// TIA Portal project "YDSLK_HMI_2023-05-10_08-26_V3_00T" (V15.1) (continued)
   "ST_HMI_Var_HMI_r64PositiveAccel_ZouChe_ChuChe" : LReal = PLC ST_HMI_Var.HMI_r64PositiveAccel_ZouChe_ChuChe AT 10-30-00-01-00-21-84-00-13-00, 1 s
   "ST_HMI_Var_HMI_r64AccVelocity_Jog_ChengXing_Up" : LReal = PLC ST_HMI_Var.HMI_r64AccVelocity_Jog_ChengXing_Up AT 10-30-00-01-00-21-84-00-1D-40, 1 s
   "VBS_time_hour" : LReal, internal
   "ST_HMI_Var_HMI_r64Velocity_Jog_JinChe" : LReal = PLC ST_HMI_Var.HMI_r64Velocity_Jog_JinChe AT 10-30-00-01-00-21-84-00-1A-40, 1 s
   "ST_HMI_Var_HMI_alpha_JuanRao_3" : LReal = PLC ST_HMI_Var.HMI_alpha_JuanRao_3 AT 10-30-00-01-00-21-84-00-33-80, 1 s
   "ST_HMI_Var_HMI_r64_LuoSha_Force_DanSha_ZhangLi_FangKai" : LReal = PLC ST_HMI_Var.HMI_r64_LuoSha_Force_DanSha_ZhangLi_FangKai AT 10-30-00-01-00-21-84-00-21-80, 1 s
   "ST_HMI_Var_HMI_r64Height_ShaSui_Start" : LReal = PLC ST_HMI_Var.HMI_r64Height_ShaSui_Start AT 10-30-00-01-00-21-84-00-0A-80, 1 s
   "ST_HMI_Var_HMI_r64Axis_ChengXing_positiveaccelstartjerk_CunRao" : LReal = PLC ST_HMI_Var.HMI_r64Axis_ChengXing_positiveaccelstartjerk_CunRao AT 10-30-00-01-00-21-84-00-3C-80, 1 s
   "ST_HMI_Var_HMI_K_T_M" : LReal = PLC ST_HMI_Var.HMI_K_T_M AT 10-30-00-01-00-21-84-00-43-C0, 1 s
   "ST_HMI_Var_HMI_r64Diameter_ShaGuan_Bottom" : LReal = PLC ST_HMI_Var.HMI_r64Diameter_ShaGuan_Bottom AT 10-30-00-01-00-21-84-00-0C-80, 1 s
   "ST_HMI_Var_HMI_r64Axis_1_ZhangLi_Position_JuanRao_Set_ND" : LReal = PLC ST_HMI_Var.HMI_r64Axis_1_ZhangLi_Position_JuanRao_Set_ND AT 10-30-00-01-00-21-84-00-39-00, 1 s
   "ST_HMI_Var_HMI_r64AccVelocity_Jog_ChuChe" : LReal = PLC ST_HMI_Var.HMI_r64AccVelocity_Jog_ChuChe AT 10-30-00-01-00-21-84-00-1A-00, 1 s
   "ST_HMI_Var_HMI_r64Velocity_Jog_ChengXing_Up" : LReal = PLC ST_HMI_Var.HMI_r64Velocity_Jog_ChengXing_Up AT 10-30-00-01-00-21-84-00-1D-00, 1 s
   "ST_HMI_Var_HMI_cam2_ratio_delt_min" : LReal = PLC ST_HMI_Var.HMI_cam2_ratio_delt_min AT 10-30-00-01-00-21-84-00-30-00, 1 s
   "ST_HMI_Var_HMI_r64Axis_DingZi_Velocity_JuanRao_max" : LReal = PLC ST_HMI_Var.HMI_r64Axis_DingZi_Velocity_JuanRao_max AT 10-30-00-01-00-21-84-00-38-40, 1 s
   "ST_Main_Var_g_bo_Automatic_Running_Status" : Bool = PLC ST_Main_Var.g_bo_Automatic_Running_Status AT 10-01-00-01-00-23-84-00-51-E0, 1 s
   "ST_HMI_Var_HMI_cam_ChengXing_delt_syncoffpositionslave_tuirao" : LReal = PLC ST_HMI_Var.HMI_cam_ChengXing_delt_syncoffpositionslave_tuirao AT 10-30-00-01-00-21-84-00-32-40, 1 s
   "变量_4" : UInt, internal
   "ST_Main_Var_g_r64Axis_DingZi_Velocity_CunRao_ratio" : LReal = PLC ST_Main_Var.g_r64Axis_DingZi_Velocity_CunRao_ratio AT 10-30-00-01-00-23-84-00-32-C0, 1 s
   "变量_2" : WString[10], internal
   "ST_HMI_Var_HMI_r64Axis_ZouChe_negativeaccelstartjerk_JinChe" : LReal = PLC ST_HMI_Var.HMI_r64Axis_ZouChe_negativeaccelstartjerk_JinChe AT 10-30-00-01-00-21-84-00-15-40, 1 s
   "ST_HMI_Var_HMI_r64Axis_1_ZhangLi_Velocity_JuanRao" : LReal = PLC ST_HMI_Var.HMI_r64Axis_1_ZhangLi_Velocity_JuanRao AT 10-30-00-01-00-21-84-00-3B-40, 1 s
   "变量_16" : Bool, internal
   "ST_HMI_Var_HMI_r64_MaoZhou_TouShu" : Int = PLC ST_HMI_Var.HMI_r64_MaoZhou_TouShu AT 10-05-00-01-00-21-84-00-22-00, 1 s
   "ST_HMI_Var_HMI_xit_delt_max" : LReal = PLC ST_HMI_Var.HMI_xit_delt_max AT 10-30-00-01-00-21-84-00-24-00, 1 s
   "ST_HMI_Var_luoshu" : Int = PLC ST_HMI_Var.luoshu AT 10-05-00-01-00-21-84-00-6B-00, 1 s
   "ST_HMI_Var_HMI_r64NianSu_3" : LReal = PLC ST_HMI_Var.HMI_r64NianSu_3 AT 10-30-00-01-00-21-84-00-04-00, 1 s
   "ST_HMI_Var_HMI_boAlarm_NianSuo_PosNon" : Bool = PLC ST_HMI_Var.HMI_boAlarm_NianSuo_PosNon AT 10-01-00-01-00-21-84-00-05-C0, 1 s
   "ST_HMI_Var_HMI_r64NianDu_actual" : LReal = PLC ST_HMI_Var.HMI_r64NianDu_actual AT 10-30-00-01-00-21-84-00-19-40, 1 s
   "ST_HMI_Var_HMI_r64Axis_ZouChe_positiveaccelendjerk_JinChe" : LReal = PLC ST_HMI_Var.HMI_r64Axis_ZouChe_positiveaccelendjerk_JinChe AT 10-30-00-01-00-21-84-00-15-00, 1 s
   "Axis_ZouChe_motionStateData_commandVelocity" : LReal = PLC Axis_ZouChe.motionStateData.commandVelocity AT A1-30-00-08-00-0A-00-00-00-6A, 1 s   // Set velocity of the axis
   "ST_Main_Var_g_bo_Mode_Enabled_Manual" : Bool = PLC ST_Main_Var.g_bo_Mode_Enabled_Manual AT 10-01-00-01-00-00-82-00-00-5A, 1 s
   "变量_8" : UInt, internal
   "ST_HMI_Var_HMI_r64_cam_ChengXing_velocity_tuirao" : LReal = PLC ST_HMI_Var.HMI_r64_cam_ChengXing_velocity_tuirao AT 10-30-00-01-00-21-84-00-30-80, 1 s
   "ST_HMI_Var_HMI_Bo_Feed_On_Off_Select" : Bool = PLC ST_HMI_Var.HMI_Bo_Feed_On_Off_Select AT 10-01-00-01-00-21-84-00-65-C0, 1 s
   "ST_HMI_Var_HMI_r64Time_TuiRao" : LReal = PLC ST_HMI_Var.HMI_r64Time_TuiRao AT 10-30-00-01-00-21-84-00-10-00, 1 s
   "ST_HMI_Var_HMI_bo_JuanRao" : Bool = PLC ST_HMI_Var.HMI_bo_JuanRao AT 10-01-00-01-00-21-84-00-6C-08, 1 s
   "ST_Main_Var_g_r64Axis_DingZi_Velocity_CunRao" : LReal = PLC ST_Main_Var.g_r64Axis_DingZi_Velocity_CunRao AT 10-30-00-01-00-23-84-00-65-C0, 1 s
   "ST_HMI_Var_HMI_r64_cam_ChengXing_positiveaccel_juanrao" : LReal = PLC ST_HMI_Var.HMI_r64_cam_ChengXing_positiveaccel_juanrao AT 10-30-00-01-00-21-84-00-36-40, 1 s
   "ST_HMI_Var_HMI_Y_L_0" : LReal = PLC ST_HMI_Var.HMI_Y_L_0 AT 10-30-00-01-00-21-84-00-42-C0, 1 s
   "变量_10" : UInt, internal
   "ST_HMI_Var_HMI_cam2_ratio_delt_ratio" : LReal = PLC ST_HMI_Var.HMI_cam2_ratio_delt_ratio AT 10-30-00-01-00-21-84-00-2F-C0, 1 s
   "ST_HMI_Var_HMI_r64QianShen_FirstArea" : LReal = PLC ST_HMI_Var.HMI_r64QianShen_FirstArea AT 10-30-00-01-00-21-84-00-07-C0, 1 s
   "ST_Cam5_Data_Var_g_ratioV" : LReal = PLC ST_Cam5_Data_Var.g_ratioV AT 10-30-00-01-00-17-84-00-01-C0, 1 s
   "ST_HMI_Var_HMI_r64_Position_DingZi_tuirao_cam2_nn_ratio_0" : LReal = PLC ST_HMI_Var.HMI_r64_Position_DingZi_tuirao_cam2_nn_ratio_0 AT 10-30-00-01-00-21-84-00-2F-00, 1 s
   "ST_HMI_Var_HMI_r64Velocity_Jog_ZhangLi_Up" : LReal = PLC ST_HMI_Var.HMI_r64Velocity_Jog_ZhangLi_Up AT 10-30-00-01-00-21-84-00-1F-C0, 1 s
   "ST_MotionTask_cam5_Comb{15}" : LReal = PLC ST_MotionTask_cam5.Comb[15] AT 10-30-00-01-00-26-84-00-0E-00, 1 s
   "VBS_maintenanceWarnStatus_8" : UInt, internal
   "ST_HMI_Var_HMI_cam2_ratio_max" : LReal = PLC ST_HMI_Var.HMI_cam2_ratio_max AT 10-30-00-01-00-21-84-00-2F-80, 1 s
   "ST_HMI_Var_HMI_r64Axis_DingZi_positiveaccelstartjerk_TuiRao" : LReal = PLC ST_HMI_Var.HMI_r64Axis_DingZi_positiveaccelstartjerk_TuiRao AT 10-30-00-01-00-21-84-00-2D-C0, 1 s
   "ST_Cam5_Data_Var_tz3" : LReal = PLC ST_Cam5_Data_Var.tz3 AT 10-30-00-01-00-17-84-00-03-00, 1 s
   "Axis_1_ZhangLi_torqueLimitPositive_value" : LReal = PLC Axis_1_ZhangLi.torqueLimitPositive.value AT A1-30-00-08-00-0B-00-00-01-2C, 1 s   // Torque limiting for the drive
   "VBS_j_times_8" : UInt, internal
   "ST_Main_Var_Axis_ChengXing_Mode_Status" : Int = PLC ST_Main_Var.Axis_ChengXing_Mode_Status AT 10-05-00-01-00-23-84-00-58-C0, 1 s
   "ST_HMI_Var_HMI_r64_cam_DingZi_negativeaccel_TuiRao" : LReal = PLC ST_HMI_Var.HMI_r64_cam_DingZi_negativeaccel_TuiRao AT 10-30-00-01-00-21-84-00-2B-80, 1 s
   "ST_HMI_Var_HMI_g1_n_delt_new_0" : LReal = PLC ST_HMI_Var.HMI_g1_n_delt_new_0 AT 10-30-00-01-00-21-84-00-39-C0, 1 s
   "ST_HMI_Var_HMI_r64NianDu_all" : LReal = PLC ST_HMI_Var.HMI_r64NianDu_all AT 10-30-00-01-00-21-84-00-01-00, 1 s
   "ST_HMI_Var_HMI_GAM_T_Z_max" : LReal = PLC ST_HMI_Var.HMI_GAM_T_Z_max AT 10-30-00-01-00-21-84-00-44-00, 1 s
   "ST_HMI_Var_HMI_r64_Lcr" : LReal = PLC ST_HMI_Var.HMI_r64_Lcr AT 10-30-00-01-00-21-84-00-3D-80, 1 s
   "ST_Main_Var_g_u32_N_Cycle_Whole" : UDInt = PLC ST_Main_Var.g_u32_N_Cycle_Whole AT 10-06-00-01-00-23-84-00-00-40, 1 s
   "ST_HMI_Var_HMI_r64Length_JuanRao" : LReal = PLC ST_HMI_Var.HMI_r64Length_JuanRao AT 10-30-00-01-00-21-84-00-05-80, 1 s
   "Axis_ZC_FU_positioningState_actualPosition" : LReal = PLC Axis_ZC_FU.positioningState.actualPosition AT A1-30-00-08-00-1D-00-00-02-23, 1 s   // Actual position of axis
   "ST_HMI_Var_HMI_r64QianShen_FenSan_real_ShengTou" : LReal = PLC ST_HMI_Var.HMI_r64QianShen_FenSan_real_ShengTou AT 10-30-00-01-00-21-84-00-71-40, 1 s
   "ST_HMI_Var_HMI_r64NianDu_1" : LReal = PLC ST_HMI_Var.HMI_r64NianDu_1 AT 10-30-00-01-00-21-84-00-02-00, 1 s
   "ST_Main_Var_ST_LuoLaSwitch" : Bool = PLC ST_Main_Var.ST_LuoLaSwitch AT 10-01-00-01-00-23-84-00-34-30, 1 s
   "ST_FC_Var_g_f1_n_piantiao_min" : LReal = PLC ST_FC_Var.g_f1_n_piantiao_min AT 10-30-00-01-00-1F-84-04-EB-80, 1 s
   "变量_25" : Int, internal
   "ST_HMI_Var_HMI_r64Axis_DingZi_Velocity_real" : LReal = PLC ST_HMI_Var.HMI_r64Axis_1_ZhangLi_PositiveAccel_from_ChengXing_ratio_tuirao AT 10-30-00-01-00-21-84-00-6E-40, 100 ms
   "ST_HMI_Var_HMI_r64_cam_ChengXing_positiveaccelstartjerk_juanrao" : LReal = PLC ST_HMI_Var.HMI_r64_cam_ChengXing_positiveaccelstartjerk_juanrao AT 10-30-00-01-00-21-84-00-36-C0, 1 s
   "ST_HMI_Var_HMI_r64Axis_1_ZhangLi_Additive_Torque_JuanRao" : LReal = PLC ST_HMI_Var.HMI_r64Axis_1_ZhangLi_Additive_Torque_JuanRao AT 10-30-00-01-00-21-84-00-3B-C0, 1 s
   "ST_FC_Var_g_f1_n_delt_ratio" : LReal = PLC ST_FC_Var.g_f1_n_delt_ratio AT 10-30-00-01-00-1F-84-04-ED-40, 1 s
   "ST_Main_Var_g_r64Axis_LuoLa_Position" : LReal = PLC ST_Main_Var.g_r64Axis_LuoLa_Position AT 10-30-00-01-00-23-84-00-1C-C0, 1 s
   "ST_HMI_Var_HMI_r64NianDu_2" : LReal = PLC ST_HMI_Var.HMI_r64NianDu_2 AT 10-30-00-01-00-21-84-00-02-40, 1 s
   "ST_HMI_Var_HMI_r64_cam_ChengXing_negativeaccelstartjerk_juanrao" : LReal = PLC ST_HMI_Var.HMI_r64_cam_ChengXing_negativeaccelstartjerk_juanrao AT 10-30-00-01-00-21-84-00-37-40, 1 s
   "ST_HMI_Var_HMI_r64_ZiDongTingZhi_NianDu_SheDing" : LReal = PLC ST_HMI_Var.HMI_r64_ZiDongTingZhi_NianDu_SheDing AT 10-30-00-01-00-21-84-00-40-C0, 1 s
   "ST_HMI_Var_HMI_r64_cam_ChengXing_negativeaccelstartjerk_tuirao" : LReal = PLC ST_HMI_Var.HMI_r64_cam_ChengXing_negativeaccelstartjerk_tuirao AT 10-30-00-01-00-21-84-00-31-C0, 1 s
   "VBS_time_day" : LReal, internal
   "变量_23" : Int, internal
   "ST_HMI_Var_HMI_r64Axis_ChengXing_positiveaccelstartjerk_TuiRao" : LReal = PLC ST_HMI_Var.HMI_r64Axis_ChengXing_positiveaccelstartjerk_TuiRao AT 10-30-00-01-00-21-84-00-26-80, 1 s
   "变量_30" : Int, internal
   "ST_HMI_Var_HMI_r64Axis_DingZi_negativeaccelendjerk_JiaNian" : LReal = PLC ST_HMI_Var.HMI_r64Axis_DingZi_negativeaccelendjerk_JiaNian AT 10-30-00-01-00-21-84-00-25-C0, 1 s
   "ST_HMI_Var_HMI_boAlarm_NianSuo_SuDuOver" : Bool = PLC ST_HMI_Var.HMI_boAlarm_NianSuo_SuDuOver AT 10-01-00-01-00-21-84-00-05-C8, 1 s
   "ST_HMI_Var_HMI_r64QianShen_All" : LReal = PLC ST_HMI_Var.HMI_r64QianShen_All AT 10-30-00-01-00-21-84-00-06-00, 1 s
   "ST_HMI_Var_HMI_r64AccVelocity_Jog_JiaNian" : LReal = PLC ST_HMI_Var.HMI_r64AccVelocity_Jog_JiaNian AT 10-30-00-01-00-21-84-00-1B-C0, 1 s
   "ST_HMI_Var_HMI_r64Axis_ChengXing_positiveaccelendjerk_TuiRao" : LReal = PLC ST_HMI_Var.HMI_r64Axis_ChengXing_positiveaccelendjerk_TuiRao AT 10-30-00-01-00-21-84-00-26-C0, 1 s
   "ST_HMI_Var_HMI_bo_LuoShaShengTou" : Bool = PLC ST_HMI_Var.HMI_bo_LuoShaShengTou AT 10-01-00-01-00-21-84-00-6C-A8, 1 s
   "ST_Main_Var_g_bo_Mode_Enabled_KongDing" : Bool = PLC ST_Main_Var.g_bo_Mode_Enabled_KongDing AT 10-01-00-01-00-00-82-00-00-51, 1 s
   "ST_HMI_Var_HMI_bo_KongDingShengTou" : Bool = PLC ST_HMI_Var.HMI_bo_KongDingShengTou AT 10-01-00-01-00-21-84-00-6C-28, 1 s
   "ST_HMI_Var_HMI_r64_DanSha_ZhangLi_ShengTou" : LReal = PLC ST_HMI_Var.HMI_r64_DanSha_ZhangLi_ShengTou AT 10-30-00-01-00-21-84-00-44-80, 1 s
   "ST_HMI_Var_HMI_r64Axis_1_ZhangLi_Position_JuanRao_Set_KongDing_12" : LReal = PLC ST_HMI_Var.HMI_r64Axis_1_ZhangLi_Position_JuanRao_Set_KongDing_12 AT 10-30-00-01-00-21-84-00-58-00, 1 s
   "Axis_LuoLa_positioningState_commandPosition" : LReal = PLC Axis_LuoLa.positioningState.commandPosition AT A1-30-00-08-00-11-00-00-02-24, 1 s
   "ST_HMI_Var_HMI_i16_QianShen_Select" : Int = PLC ST_HMI_Var.HMI_i16_QianShen_Select AT 10-05-00-01-00-21-84-00-08-90, 1 s
   "ST_HMI_Var_HMI_r64NegativeAccel_ZouChe_ChuChe" : LReal = PLC ST_HMI_Var.HMI_r64NegativeAccel_ZouChe_ChuChe AT 10-30-00-01-00-21-84-00-13-40, 1 s
   "ST_HMI_Var_HMI_r64Axis_ZouChe_Position_KongDing_8" : LReal = PLC ST_HMI_Var.HMI_r64Axis_ZouChe_Position_KongDing_8 AT 10-30-00-01-00-21-84-00-50-00, 1 s
   "ST_HMI_Var_HMI_r64Axis_ChengXing_Position_delt_KongDing_8" : LReal = PLC ST_HMI_Var.HMI_r64Axis_ChengXing_Position_delt_KongDing_8 AT 10-30-00-01-00-21-84-00-51-40, 1 s
   "ST_HMI_Var_HMI_r64_DingZi_Zouche_ratio_KongDing_9" : LReal = PLC ST_HMI_Var.HMI_r64_DingZi_Zouche_ratio_KongDing_9 AT 10-30-00-01-00-21-84-00-52-C0, 1 s
   "ST_HMI_Var_HMI_r64Axis_ZouChe_Position_LuoSha_8" : LReal = PLC ST_HMI_Var.HMI_r64Axis_ZouChe_Position_LuoSha_8 AT 10-30-00-01-00-21-84-00-5D-C0, 1 s
   "ST_HMI_Var_HMI_r64_DingZi_Zouche_ratio_LuoSha_9" : LReal = PLC ST_HMI_Var.HMI_r64_DingZi_Zouche_ratio_LuoSha_9 AT 10-30-00-01-00-21-84-00-60-C0, 1 s
   "ST_HMI_Var_HMI_r64Axis_ZouChe_Position_KongDing_9" : LReal = PLC ST_HMI_Var.HMI_r64Axis_ZouChe_Position_KongDing_9 AT 10-30-00-01-00-21-84-00-51-C0, 1 s
   "ST_HMI_Var_HMI_r64Axis_1_ZhangLi_Position_JuanRao_real2" : Int = PLC ST_HMI_Var.HMI_r64Axis_1_ZhangLi_Position_JuanRao_real2 AT 10-05-00-01-00-21-84-00-6F-80, 100 ms
   "ST_HMI_Var_HMI_r64Axis_ChengXing_Position_real2" : Int = PLC ST_HMI_Var.HMI_r64Axis_ChengXing_Position_real2 AT 10-05-00-01-00-21-84-00-70-40, 1 s
   "ST_HMI_Var_HMI_r64Axis_ZouChe_Position_real" : LReal = PLC ST_HMI_Var.HMI_r64Axis_ZouChe_Position_real AT 10-30-00-01-00-21-84-00-6D-40, 100 ms
   "ST_HMI_Var_HMI_r64Axis_ZouChe_Position_real2" : Int = PLC ST_HMI_Var.HMI_r64Axis_ZouChe_Position_real2 AT 10-05-00-01-00-21-84-00-6D-80, 100 ms
   "ST_Main_Var_g_u16_N_Cycle_Single(1)" : UInt = PLC ST_Main_Var.g_u16_N_Cycle_Single AT 10-04-00-01-00-23-84-00-00-10, 1 s
   "ST_FC_Var_g_N" : LReal = PLC ST_FC_Var.g_N AT 10-30-00-01-00-1F-84-00-0D-40, 1 s
   "ST_FC_Var_g_ND" : LReal = PLC ST_FC_Var.g_ND AT 10-30-00-01-00-1F-84-00-0C-C0, 1 s
   "VBS_hengsi_status0" : Int, internal
   "VBS_hengsi_status1" : Int, internal
   "ST_HMI_Var_HMI_i16_ShengTou_Select" : Int = PLC ST_HMI_Var.HMI_i16_ShengTou_Select AT 10-05-00-01-00-21-84-00-72-10, 1 s
   "ST_Main_Var_g_bo_KongDing_Running_Status" : Bool = PLC ST_Main_Var.g_bo_KongDing_Running_Status AT 10-01-00-01-00-23-84-00-57-B0, 1 s
   "ST_HMI_Var_HMI_r64Axis_ChengXing_Position_real" : LReal = PLC ST_HMI_Var.HMI_r64Axis_ChengXing_Position_real AT 10-30-00-01-00-21-84-00-70-00, 1 s
   "ST_Main_Var_g_bo_ZiDong_JiTing" : Bool = PLC ST_Main_Var.g_bo_ZiDong_JiTing AT 10-01-00-01-00-00-81-00-00-28, 1 s
   "ST_Main_Var_g_SLM_enable_status" : Bool = PLC ST_Main_Var.g_SLM_enable_status AT 10-01-00-01-00-23-84-00-59-B0, 1 s
   "ST_HMI_Var_HMI_bo_Auto" : Bool = PLC ST_HMI_Var.HMI_bo_Auto AT 10-01-00-01-00-21-84-00-6C-48, 1 s
   "ST_HMI_Var_HMI_r64QianShen_All_KongDing_7" : LReal = PLC ST_HMI_Var.HMI_r64QianShen_All_KongDing_7 AT 10-30-00-01-00-21-84-00-4D-C0, 1 s
   "ST_HMI_Var_HMI_r64QianShen_FenSan_KongDing_7" : LReal = PLC ST_HMI_Var.HMI_r64QianShen_FenSan_KongDing_7 AT 10-30-00-01-00-21-84-00-4E-00, 1 s
   "ST_HMI_Var_HMI_bo_QianShen_ShengTou_Add" : Bool = PLC ST_HMI_Var.HMI_bo_QianShen_ShengTou_Add AT 10-01-00-01-00-21-84-00-71-80, 1 s
   "ST_HMI_Var_HMI_bo_QianShen_ShengTou_Minus" : Bool = PLC ST_HMI_Var.HMI_bo_QianShen_ShengTou_Minus AT 10-01-00-01-00-21-84-00-71-88, 1 s
   "ST_HMI_Var_HMI_r64NianDu_QianShen_Best" : LReal = PLC ST_HMI_Var.HMI_r64NianDu_QianShen_Best AT 10-30-00-01-00-21-84-00-01-40, 1 s
   "ST_HMI_Var_HMI_r64_Scale_KongDing_7" : LReal = PLC ST_HMI_Var.HMI_r64_Scale_KongDing_7 AT 10-30-00-01-00-21-84-00-4E-40, 1 s
   "ST_HMI_Var_HMI_r64Position_ChuChe_KongDing_7" : LReal = PLC ST_HMI_Var.HMI_r64Position_ChuChe_KongDing_7 AT 10-30-00-01-00-21-84-00-4D-80, 1 s
   "ST_HMI_Var_HMI_r64QianShen_First_UpperLimit" : LReal = PLC ST_HMI_Var.HMI_r64QianShen_First_UpperLimit AT 10-30-00-01-00-21-84-00-07-80, 1 s
   "ST_HMI_Var_HMI_r64StartPosition_Axis_ZouChe_0" : LReal = PLC ST_HMI_Var.HMI_r64StartPosition_Axis_ZouChe_0 AT 10-30-00-01-00-21-84-00-18-40, 1 s
   "ST_HMI_Var_HMI_r64StartPosition_Axis_1_ZhangLi_0" : LReal = PLC ST_HMI_Var.HMI_r64StartPosition_Axis_1_ZhangLi_0 AT 10-30-00-01-00-21-84-00-18-C0, 1 s
   "ST_HMI_Var_HMI_r64StartPosition_Axis_ChengXing_0" : LReal = PLC ST_HMI_Var.HMI_r64StartPosition_Axis_ChengXing_0 AT 10-30-00-01-00-21-84-00-18-80, 1 s
   "Axis_2_ZhangLi_positioningState_actualPosition" : LReal = PLC Axis_2_ZhangLi.positioningState.actualPosition AT A1-30-00-08-00-19-00-00-02-23, 1 s
   "Axis_1_ZhangLi_positioningState_actualPosition" : LReal = PLC Axis_1_ZhangLi.positioningState.actualPosition AT A1-30-00-08-00-0B-00-00-02-23, 1 s
   "Axis_ChengXing_positioningState_actualPosition" : LReal = PLC Axis_ChengXing.positioningState.actualPosition AT A1-30-00-08-00-0C-00-00-02-23, 1 s
   "ST_HMI_Var_HMI_boMinorAdjustment_select" : Bool = PLC ST_HMI_Var.HMI_boMinorAdjustment_select AT 10-01-00-01-00-21-84-00-19-80, 1 s
   "ST_Var_ZLCD_HMI_r64Axis_1_ZhangLi_Position_CeDing_N{0}" : LReal = PLC ST_Var_ZLCD.HMI_r64Axis_1_ZhangLi_Position_CeDing_N[0] AT 10-30-00-01-00-34-84-00-01-80, 1 s
   "ST_Var_ZLCD_HMI_r64Axis_1_ZhangLi_Torque_CeDing_N{0}" : LReal = PLC ST_Var_ZLCD.HMI_r64Axis_1_ZhangLi_Torque_CeDing_N[0] AT 10-30-00-01-00-34-84-00-29-C0, 1 s
   "ST_Var_ZLCD_HMI_r64Axis_1_ZhangLi_Torque_CeDing_N{1}" : LReal = PLC ST_Var_ZLCD.HMI_r64Axis_1_ZhangLi_Torque_CeDing_N[1] AT 10-30-00-01-00-34-84-00-2A-00, 1 s
   "ST_Var_ZLCD_HMI_r64Axis_1_ZhangLi_Torque_CeDing_N{2}" : LReal = PLC ST_Var_ZLCD.HMI_r64Axis_1_ZhangLi_Torque_CeDing_N[2] AT 10-30-00-01-00-34-84-00-2A-40, 1 s
   "ST_Var_ZLCD_HMI_r64Axis_1_ZhangLi_Torque_CeDing_N{3}" : LReal = PLC ST_Var_ZLCD.HMI_r64Axis_1_ZhangLi_Torque_CeDing_N[3] AT 10-30-00-01-00-34-84-00-2A-80, 1 s
   "ST_Var_ZLCD_HMI_r64Axis_1_ZhangLi_Torque_CeDing_N{4}" : LReal = PLC ST_Var_ZLCD.HMI_r64Axis_1_ZhangLi_Torque_CeDing_N[4] AT 10-30-00-01-00-34-84-00-2A-C0, 1 s
   "ST_Var_ZLCD_HMI_r64Axis_1_ZhangLi_Torque_CeDing_N{6}" : LReal = PLC ST_Var_ZLCD.HMI_r64Axis_1_ZhangLi_Torque_CeDing_N[6] AT 10-30-00-01-00-34-84-00-2B-40, 1 s
   "ST_Var_ZLCD_HMI_bo_ZhangLi_CeDing_Adjustment" : Bool = PLC ST_Var_ZLCD.HMI_bo_ZhangLi_CeDing_Adjustment AT 10-01-00-01-00-34-84-00-01-40, 1 s
   "ST_HMI_Var_HMI_r64_h0_s" : LReal = PLC ST_HMI_Var.HMI_r64_h0_s AT 10-30-00-01-00-21-84-00-0D-40, 1 s
   "ST_HMI_Var_HMI_r64Axis_ZouChe_Position_LuoSha_9" : LReal = PLC ST_HMI_Var.HMI_r64Axis_ZouChe_Position_LuoSha_9 AT 10-30-00-01-00-21-84-00-60-80, 1 s
   "ST_HMI_Var_HMI_r64Position_ChuChe_KongDing_65" : LReal = PLC ST_HMI_Var.HMI_r64Position_ChuChe_KongDing_65 AT 10-30-00-01-00-21-84-00-4C-80, 1 s
   "ST_HMI_Var_HMI_r64QianShen_KongDing_65" : LReal = PLC ST_HMI_Var.HMI_r64QianShen_KongDing_65 AT 10-30-00-01-00-21-84-00-4C-C0, 1 s
   "ST_HMI_Var_HMI_r64_DingZi_Zouche_ratio_KongDing_65" : LReal = PLC ST_HMI_Var.HMI_r64_DingZi_Zouche_ratio_KongDing_65 AT 10-30-00-01-00-21-84-00-4D-00, 1 s
   "ST_Main_Var_g_i16_KongDing_Status" : Int = PLC ST_Main_Var.g_i16_KongDing_Status AT 10-05-00-01-00-23-84-00-55-F0, 1 s
   "ST_HMI_Var_HMI_r64NianSu_Max" : LReal = PLC ST_HMI_Var.HMI_r64NianSu_Max AT 10-30-00-01-00-21-84-00-04-40, 1 s
   "ST_HMI_Var_HMI_r64Ratio_PositiveAccel_Jerk_JiaNian" : LReal = PLC ST_HMI_Var.HMI_r64Ratio_PositiveAccel_Jerk_JiaNian AT 10-30-00-01-00-21-84-00-01-80, 1 s
   "ST_Calculation_Var_g_r64Axis_DingZi_PositiveAccel_Buffer_JiaNian{0}" : LReal = PLC ST_Calculation_Var.g_r64Axis_DingZi_PositiveAccel_Buffer_JiaNian[0] AT 10-30-00-01-00-13-84-00-0D-40, 1 s
   "ST_Calculation_Var_Date_Temp" : Int = PLC ST_Calculation_Var.Date_Temp AT 10-05-00-01-00-13-84-00-00-90, 1 s
   "ST_Calculation_Var_g_r64Axis_DingZi_PositiveAccel_Buffer_JiaNian{1}" : LReal = PLC ST_Calculation_Var.g_r64Axis_DingZi_PositiveAccel_Buffer_JiaNian[1] AT 10-30-00-01-00-13-84-00-0D-80, 1 s
   "ST_Calculation_Var_g_r64Axis_DingZi_PositiveAccelStartJerk_Buffer_JiaNian{0}" : LReal = PLC ST_Calculation_Var.g_r64Axis_DingZi_PositiveAccelStartJerk_Buffer_JiaNian[0] AT 10-30-00-01-00-13-84-00-0E-40, 1 s
   "ST_Calculation_Var_g_r64Axis_DingZi_PositiveAccelStartJerk_Buffer_JiaNian{1}" : LReal = PLC ST_Calculation_Var.g_r64Axis_DingZi_PositiveAccelStartJerk_Buffer_JiaNian[1] AT 10-30-00-01-00-13-84-00-0E-80, 1 s
   "ST_HMI_Var_HMI_i16_Status_ShaGuan_Select" : Int = PLC ST_HMI_Var.HMI_i16_Status_ShaGuan_Select AT 10-05-00-01-00-21-84-00-0C-40, 1 s
   "ST_HMI_Var_HMI_r64Diameter_ShaGuan_Bottom_2" : LReal = PLC ST_HMI_Var.HMI_r64Diameter_ShaGuan_Bottom_2 AT 10-30-00-01-00-21-84-00-0E-00, 1 s
   "ST_HMI_Var_HMI_r64_h0_s_2" : LReal = PLC ST_HMI_Var.HMI_r64_h0_s_2 AT 10-30-00-01-00-21-84-00-0E-C0, 1 s
   "ST_HMI_Var_HMI_r64Diameter_ShaGuan_Middle_2" : LReal = PLC ST_HMI_Var.HMI_r64Diameter_ShaGuan_Middle_2 AT 10-30-00-01-00-21-84-00-0E-40, 1 s
   "ST_HMI_Var_HMI_r64Diameter_ShaGuan_Top_2" : LReal = PLC ST_HMI_Var.HMI_r64Diameter_ShaGuan_Top_2 AT 10-30-00-01-00-21-84-00-0E-80, 1 s
   "ST_HMI_Var_HMI_r64Height_ShaGuan_Middle_2" : LReal = PLC ST_HMI_Var.HMI_r64Height_ShaGuan_Middle_2 AT 10-30-00-01-00-21-84-00-0F-00, 1 s
   "ST_HMI_Var_HMI_r64Height_ShaGuan_Top_2" : LReal = PLC ST_HMI_Var.HMI_r64Height_ShaGuan_Top_2 AT 10-30-00-01-00-21-84-00-0F-40, 1 s
   "ST_HMI_Var_HMI_r64Axis_ZouChe_Position_ShengTou_Start_Position" : LReal = PLC ST_HMI_Var.HMI_r64Axis_ZouChe_Position_ShengTou_Start_Position AT 10-30-00-01-00-21-84-00-44-40, 1 s
   "ST_HMI_Var_HMI_bo_KongDingShengTou_GuangDing" : Bool = PLC ST_HMI_Var.HMI_bo_KongDingShengTou_GuangDing AT 10-01-00-01-00-21-84-00-6C-30, 1 s
   "ST_HMI_Var_HMI_r64Axis_ZouChe_Position_KongDing_8_1" : LReal = PLC ST_HMI_Var.HMI_r64Axis_ZouChe_Position_KongDing_8_1 AT 10-30-00-01-00-21-84-00-50-40, 1 s
   "ST_HMI_Var_HMI_r64_DingZi_Zouche_ratio_KongDing_9_1" : LReal = PLC ST_HMI_Var.HMI_r64_DingZi_Zouche_ratio_KongDing_9_1 AT 10-30-00-01-00-21-84-00-53-80, 1 s
   "Axis_ZouChe_motionStateData_actualVelocity" : LReal = PLC Axis_ZouChe.motionStateData.actualVelocity AT A1-30-00-08-00-0A-00-00-00-68, 1 s
   "HMI_Tag_bo_showDebugButton" : Bool, internal   // 显示调试画面按钮
   "Axis_LuoLa_motionStateData_actualVelocity" : LReal = PLC Axis_LuoLa.motionStateData.actualVelocity AT A1-30-00-08-00-11-00-00-00-68, 1 s
   "ST_HMI_Var_HMI_r64_DingZi_Zouche_ratio_KongDing_9_Shaguan2" : LReal = PLC ST_HMI_Var.HMI_r64_DingZi_Zouche_ratio_KongDing_9_Shaguan2 AT 10-30-00-01-00-21-84-00-53-40, 1 s
   "ST_HMI_Var_HMI_r64_DingZi_Zouche_ratio_KongDing_9_Shaguan1" : LReal = PLC ST_HMI_Var.HMI_r64_DingZi_Zouche_ratio_KongDing_9_Shaguan1 AT 10-30-00-01-00-21-84-00-53-00, 1 s
   "ST_HMI_Var_HMI_i16_Dingzi_50102AlarmStatus" : Int = PLC ST_HMI_Var.HMI_i16_Dingzi_50102AlarmStatus AT 10-05-00-01-00-21-84-00-61-D0, 1 s
   "ST_HMI_Var_HMI_bo_XiangLing" : Bool = PLC ST_HMI_Var.HMI_bo_XiangLing AT 10-01-00-01-00-21-84-00-6C-58, 1 s
   "ST_HMI_Var_HMI_i16_NianduAlarmStatus" : Int = PLC ST_HMI_Var.HMI_i16_NianduAlarmStatus AT 10-05-00-01-00-21-84-00-61-C0, 1 s
   "ST_HMI_Var_HMI_r64_QianShen_Add1" : LReal = PLC ST_HMI_Var.HMI_r64_QianShen_Add1 AT 10-30-00-01-00-21-84-00-62-00, 1 s
   "ST_HMI_Var_HMI_r64_QianShen_Add2" : LReal = PLC ST_HMI_Var.HMI_r64_QianShen_Add2 AT 10-30-00-01-00-21-84-00-62-40, 1 s
   "ST_HMI_Var_HMI_r64_ShaXian_L1" : LReal = PLC ST_HMI_Var.HMI_r64_ShaXian_L1 AT 10-30-00-01-00-21-84-00-62-80, 1 s
   "ST_HMI_Var_HMI_r64_Ratio1" : LReal = PLC ST_HMI_Var.HMI_r64_Ratio1 AT 10-30-00-01-00-21-84-00-63-40, 1 s
   "ST_HMI_Var_HMI_r64_ShaXian_L2" : LReal = PLC ST_HMI_Var.HMI_r64_ShaXian_L2 AT 10-30-00-01-00-21-84-00-62-C0, 1 s
   "ST_HMI_Var_HMI_r64_Ratio2" : LReal = PLC ST_HMI_Var.HMI_r64_Ratio2 AT 10-30-00-01-00-21-84-00-63-80, 1 s
   "ST_HMI_Var_HMI_r64QianShen_All_object" : LReal = PLC ST_HMI_Var.HMI_r64QianShen_All_object AT 10-30-00-01-00-21-84-00-65-40, 1 s
   "ST_HMI_Var_HMI_bo_DianYuan_Duan" : Bool = PLC ST_HMI_Var.HMI_bo_DianYuan_Duan AT 10-01-00-01-00-21-84-00-6C-50, 1 s
   "ST_HMI_Var_HMI_bo_ZiDong_QiDong" : Bool = PLC ST_HMI_Var.HMI_bo_ZiDong_QiDong AT 10-01-00-01-00-21-84-00-6C-80, 1 s
   "ST_HMI_Var_HMI_bo_Start_Position" : Bool = PLC ST_HMI_Var.HMI_bo_Start_Position AT 10-01-00-01-00-21-84-00-6C-38, 1 s
   "ST_HMI_Var_HMI_bo_Manual" : Bool = PLC ST_HMI_Var.HMI_bo_Manual AT 10-01-00-01-00-21-84-00-6C-20, 1 s
   "ST_HMI_Var_HMI_bo_Disable" : Bool = PLC ST_HMI_Var.HMI_bo_Disable AT 10-01-00-01-00-21-84-00-6C-40, 1 s
   "ST_HMI_Var_HMI_i32_ZouChe_ZhanJu_ss_1" : DInt = PLC ST_HMI_Var.HMI_i32_ZouChe_ZhanJu_ss_1 AT 10-07-00-01-00-21-84-00-70-60, 1 s
   "ST_Main_Var_g_bo_JianNian_Jog_Status" : Bool = PLC ST_Main_Var.g_bo_JianNian_Jog_Status AT 10-01-00-01-00-23-84-00-65-50, 1 s
   "ST_Main_Var_g_bo_DI_1_D435_X122_2" : Bool = PLC ST_Main_Var.g_bo_DI_1_D435_X122_2 AT 10-01-00-01-00-23-84-00-2C-A0, 1 s
   "ST_HMI_Var_HMI_i16_ZouChe_ZhanJu_Select" : Int = PLC ST_HMI_Var.HMI_i16_ZouChe_ZhanJu_Select AT 10-05-00-01-00-21-84-00-11-00, 1 s
   "ST_HMI_Var_HMI_bo_ZouChe_ZhanJu_Select" : Bool = PLC ST_HMI_Var.HMI_bo_ZouChe_ZhanJu_Select AT 10-01-00-01-00-21-84-00-70-50, 1 s
   "ST_HMI_Var_HMI_r64_ZouChe_ZhanJu_Max_20" : LReal = PLC ST_HMI_Var.HMI_r64_ZouChe_ZhanJu_Max_20 AT 10-30-00-01-00-21-84-00-11-80, 1 s
   "ST_HMI_Var_HMI_r64_ZouChe_ZhanJu_Max_25" : LReal = PLC ST_HMI_Var.HMI_r64_ZouChe_ZhanJu_Max_25 AT 10-30-00-01-00-21-84-00-11-C0, 1 s
   "ST_HMI_Var_HMI_r64_ZouChe_ZhanJu_Max_30" : LReal = PLC ST_HMI_Var.HMI_r64_ZouChe_ZhanJu_Max_30 AT 10-30-00-01-00-21-84-00-12-00, 1 s
   "ST_HMI_Var_HMI_r64_ZouChe_ZhanJu_Max_35" : LReal = PLC ST_HMI_Var.HMI_r64_ZouChe_ZhanJu_Max_35 AT 10-30-00-01-00-21-84-00-12-40, 1 s
   "ST_HMI_Var_HMI_r64_ZouChe_ZhanJu_Max_40" : LReal = PLC ST_HMI_Var.HMI_r64_ZouChe_ZhanJu_Max_40 AT 10-30-00-01-00-21-84-00-12-80, 1 s
   "ST_HMI_Var_HMI_r64_ZouChe_ZhanJu_Max_45" : LReal = PLC ST_HMI_Var.HMI_r64_ZouChe_ZhanJu_Max_45 AT 10-30-00-01-00-21-84-00-12-C0, 1 s
   "ST_HMI_Var_HMI_r64_ZouChe_ZhanJu_Max_Effect" : LReal = PLC ST_HMI_Var.HMI_r64_ZouChe_ZhanJu_Max_Effect AT 10-30-00-01-00-21-84-00-11-40, 1 s
   "HMI_Tag_1" : Int, internal
   "变量_100" : UInt, internal
   "ST_HMI_Var_HMI_bo_BaShaTou_Select" : Bool = PLC ST_HMI_Var.HMI_bo_BaShaTou_Select AT 10-01-00-01-00-21-84-00-72-30, 1 s
   "ST_HMI_Var_HMI_r64Axis_ZouChe_Position_LuoSha_112_Delta_BaTou" : LReal = PLC ST_HMI_Var.HMI_r64Axis_ZouChe_Position_LuoSha_112_Delta_BaTou AT 10-30-00-01-00-21-84-00-61-00, 1 s
   "ST_MotionTask_ZhangLi_Var_HMI_bo_TaiGong" : Bool = PLC ST_MotionTask_ZhangLi_Var.HMI_bo_TaiGong AT 10-01-00-01-00-25-84-00-09-D0, 1 s
   "ST_MotionTask_ZhangLi_Var_HMI_r64Axis_1_ZhangLi_Position_TaiGong" : LReal = PLC ST_MotionTask_ZhangLi_Var.HMI_r64Axis_1_ZhangLi_Position_TaiGong AT 10-30-00-01-00-25-84-00-00-C0, 1 s
   "ST_MotionTask_ZhangLi_Var_HMI_r64Axis_ZouChe_Position_TaiGong_FangXia" : LReal = PLC ST_MotionTask_ZhangLi_Var.HMI_r64Axis_ZouChe_Position_TaiGong_FangXia AT 10-30-00-01-00-25-84-00-01-80, 1 s
   "ST_Maintenance_g_u16_TimeInterval_OilChange" : UInt = PLC ST_Maintenance.g_u16_TimeInterval_OilChange AT 10-04-00-01-00-24-84-00-01-40, 1 s
   "ST_Maintenance_g_u16_TimeReminder_Maintennance" : UInt = PLC ST_Maintenance.g_u16_TimeReminder_Maintennance AT 10-04-00-01-00-24-84-00-01-50, 1 s
   "ST_Maintenance_g_u16_1_Times_OilChange_DingZi" : UInt = PLC ST_Maintenance.g_u16_1_Times_OilChange_DingZi AT 10-04-00-01-00-24-84-00-01-60, 1 s
   "ST_Maintenance_g_u16_2_Times_LongDai_HuangYouZui" : UInt = PLC ST_Maintenance.g_u16_2_Times_LongDai_HuangYouZui AT 10-04-00-01-00-24-84-00-01-70, 1 s
   "ST_Maintenance_g_u16_3_Times_LongDai_YaJinQi" : UInt = PLC ST_Maintenance.g_u16_3_Times_LongDai_YaJinQi AT 10-04-00-01-00-24-84-00-01-80, 1 s
   "ST_Maintenance_g_u16_4_Times_GongZhou_Bearing" : UInt = PLC ST_Maintenance.g_u16_4_Times_GongZhou_Bearing AT 10-04-00-01-00-24-84-00-01-90, 1 s
   "ST_Maintenance_g_u16_5_Times_LongDai_Clean" : UInt = PLC ST_Maintenance.g_u16_5_Times_LongDai_Clean AT 10-04-00-01-00-24-84-00-01-A0, 1 s
   "ST_Maintenance_g_u16_6_Times_DingZi_ChuanDong" : UInt = PLC ST_Maintenance.g_u16_6_Times_DingZi_ChuanDong AT 10-04-00-01-00-24-84-00-01-B0, 1 s
   "ST_Maintenance_g_u16_7_Times_ControlBox_Clean" : UInt = PLC ST_Maintenance.g_u16_7_Times_ControlBox_Clean AT 10-04-00-01-00-24-84-00-01-C0, 1 s
   "ST_Maintenance_g_u16_8_Times_DingZi_Fan" : UInt = PLC ST_Maintenance.g_u16_8_Times_DingZi_Fan AT 10-04-00-01-00-24-84-00-01-D0, 1 s
   "ST_Maintenance_g_u16_8_Times_TiShi_DingZi_Fan" : UInt = PLC ST_Maintenance.g_u16_8_Times_TiShi_DingZi_Fan AT 10-04-00-01-00-24-84-00-06-F0, 1 s
   "ST_Maintenance_g_bo_8_Warn_Status_DingZi_Fan" : Bool = PLC ST_Maintenance.g_bo_8_Warn_Status_DingZi_Fan AT 10-01-00-01-00-24-84-00-05-58, 1 s
   "ST_Maintenance_g_bo_8_Status_DingZi_Fan" : Bool = PLC ST_Maintenance.g_bo_8_Status_DingZi_Fan AT 10-01-00-01-00-24-84-00-05-18, 1 s
   "ST_Maintenance_g_bo_7_Warn_Status_ControlBox_Clean" : Bool = PLC ST_Maintenance.g_bo_7_Warn_Status_ControlBox_Clean AT 10-01-00-01-00-24-84-00-05-50, 1 s
   "ST_Maintenance_g_u16_7_Times_TiShi_ControlBox_Clean" : UInt = PLC ST_Maintenance.g_u16_7_Times_TiShi_ControlBox_Clean AT 10-04-00-01-00-24-84-00-06-E0, 1 s
   "ST_Maintenance_g_bo_7_Status_ControlBox_Clean" : Bool = PLC ST_Maintenance.g_bo_7_Status_ControlBox_Clean AT 10-01-00-01-00-24-84-00-05-10, 1 s
   "ST_Maintenance_g_bo_6_Warn_Status_DingZi_ChuanDong" : Bool = PLC ST_Maintenance.g_bo_6_Warn_Status_DingZi_ChuanDong AT 10-01-00-01-00-24-84-00-05-48, 1 s
   "ST_Maintenance_g_u16_6_Times_TiShi_DingZi_ChuanDong" : UInt = PLC ST_Maintenance.g_u16_6_Times_TiShi_DingZi_ChuanDong AT 10-04-00-01-00-24-84-00-06-D0, 1 s
   "ST_Maintenance_g_bo_6_Status_DingZi_ChuanDong" : Bool = PLC ST_Maintenance.g_bo_6_Status_DingZi_ChuanDong AT 10-01-00-01-00-24-84-00-05-08, 1 s
   "ST_Maintenance_g_bo_5_Warn_Status_LongDai_Clean" : Bool = PLC ST_Maintenance.g_bo_5_Warn_Status_LongDai_Clean AT 10-01-00-01-00-24-84-00-05-40, 1 s
   "ST_Maintenance_g_u16_5_Times_TiShi_LongDai_Clean" : UInt = PLC ST_Maintenance.g_u16_5_Times_TiShi_LongDai_Clean AT 10-04-00-01-00-24-84-00-06-C0, 1 s
   "ST_Maintenance_g_bo_5_Status_LongDai_Clean" : Bool = PLC ST_Maintenance.g_bo_5_Status_LongDai_Clean AT 10-01-00-01-00-24-84-00-05-00, 1 s
   "ST_Maintenance_g_bo_4_Warn_Status_GongZhou_Bearing" : Bool = PLC ST_Maintenance.g_bo_4_Warn_Status_GongZhou_Bearing AT 10-01-00-01-00-24-84-00-05-38, 1 s
   "ST_Maintenance_g_u16_4_Times_TiShi_GongZhou_Bearing" : UInt = PLC ST_Maintenance.g_u16_4_Times_TiShi_GongZhou_Bearing AT 10-04-00-01-00-24-84-00-06-B0, 1 s
   "ST_Maintenance_g_bo_4_Status_GongZhou_Bearing" : Bool = PLC ST_Maintenance.g_bo_4_Status_GongZhou_Bearing AT 10-01-00-01-00-24-84-00-04-F8, 1 s
   "ST_Maintenance_g_bo_3_Warn_Status_LongDai_YaJinQi" : Bool = PLC ST_Maintenance.g_bo_3_Warn_Status_LongDai_YaJinQi AT 10-01-00-01-00-24-84-00-05-30, 1 s
   "ST_Maintenance_g_u16_3_Times_TiShi_LongDai_YaJinQi" : UInt = PLC ST_Maintenance.g_u16_3_Times_TiShi_LongDai_YaJinQi AT 10-04-00-01-00-24-84-00-06-A0, 1 s
   "ST_Maintenance_g_bo_3_Status_LongDai_YaJinQi" : Bool = PLC ST_Maintenance.g_bo_3_Status_LongDai_YaJinQi AT 10-01-00-01-00-24-84-00-04-F0, 1 s
   "ST_Maintenance_g_bo_2_Warn_Status_LongDai_HuangYouZui" : Bool = PLC ST_Maintenance.g_bo_2_Warn_Status_LongDai_HuangYouZui AT 10-01-00-01-00-24-84-00-05-28, 1 s
   "ST_Maintenance_g_u16_2_Times_TiShi_LongDai_HuangYouZui" : UInt = PLC ST_Maintenance.g_u16_2_Times_TiShi_LongDai_HuangYouZui AT 10-04-00-01-00-24-84-00-06-90, 1 s
   "ST_Maintenance_g_bo_2_Status_LongDai_HuangYouZui" : Bool = PLC ST_Maintenance.g_bo_2_Status_LongDai_HuangYouZui AT 10-01-00-01-00-24-84-00-04-E8, 1 s
   "ST_Maintenance_g_bo_1_Warn_Status_OilChange_DingZi" : Bool = PLC ST_Maintenance.g_bo_1_Warn_Status_OilChange_DingZi AT 10-01-00-01-00-24-84-00-05-20, 1 s
   "ST_Maintenance_g_u16_1_Times_TiShi_OilChange_DingZi" : UInt = PLC ST_Maintenance.g_u16_1_Times_TiShi_OilChange_DingZi AT 10-04-00-01-00-24-84-00-06-80, 1 s
   "ST_Maintenance_g_bo_1_Status_OilChange_DingZi" : Bool = PLC ST_Maintenance.g_bo_1_Status_OilChange_DingZi AT 10-01-00-01-00-24-84-00-04-E0, 1 s
   "ST_Maintenance_g_r64_Time_All" : LReal = PLC ST_Maintenance.g_r64_Time_All AT 10-30-00-01-00-24-84-00-01-00, 1 s
   "ST_HMI_Var_HMI_r64Axis_ZouChe_Position_KongDing_12" : LReal = PLC ST_HMI_Var.HMI_r64Axis_ZouChe_Position_KongDing_12 AT 10-30-00-01-00-21-84-00-55-00, 1 s
   "ST_HMI_Var_HMI_bo_ChuChe_Middle_Select" : Bool = PLC ST_HMI_Var.HMI_bo_ChuChe_Middle_Select AT 10-01-00-01-00-21-84-00-71-90, 1 s
   "ST_HMI_Var_HMI_r64Axis_ZouChe_Position_ChuChe_Middle" : LReal = PLC ST_HMI_Var.HMI_r64Axis_ZouChe_Position_ChuChe_Middle AT 10-30-00-01-00-21-84-00-6B-40, 1 s
   "ST_Maintenance_HMI_r64_Production" : LReal = PLC ST_Maintenance.HMI_r64_Production AT 10-30-00-01-00-24-84-00-00-40, 1 s
   "ST_Maintenance_HMI_r64_Production_Once" : LReal = PLC ST_Maintenance.HMI_r64_Production_Once AT 10-30-00-01-00-24-84-00-00-80, 1 s
   "ST_Maintenance_HMI_r64_Weight_ShaSui" : LReal = PLC ST_Maintenance.HMI_r64_Weight_ShaSui AT 10-30-00-01-00-24-84-00-00-C0, 1 s
   "ST_HMI_Var_HMI_bo_ChengXing_Holding_Brake_Open" : Bool = PLC ST_HMI_Var.HMI_bo_ChengXing_Holding_Brake_Open AT 10-01-00-01-00-21-84-00-72-40, 1 s
   "ST_HMI_Var_HMI_bo_ZhangLi_Holding_Brake_Open" : Bool = PLC ST_HMI_Var.HMI_bo_ZhangLi_Holding_Brake_Open AT 10-01-00-01-00-21-84-00-72-48, 1 s
   "ST_TO_DZ_FU_Var_HMI_r64Ratio_PositiveAccelStartJerk_JiaNian" : LReal = PLC ST_TO_DZ_FU_Var.HMI_r64Ratio_PositiveAccelStartJerk_JiaNian AT 10-30-00-01-00-37-84-00-00-40, 1 s
   "ST_TO_DZ_FU_Var_HMI_r64Ratio_PositiveAccelEndJerk_JiaNian" : LReal = PLC ST_TO_DZ_FU_Var.HMI_r64Ratio_PositiveAccelEndJerk_JiaNian AT 10-30-00-01-00-37-84-00-00-80, 1 s